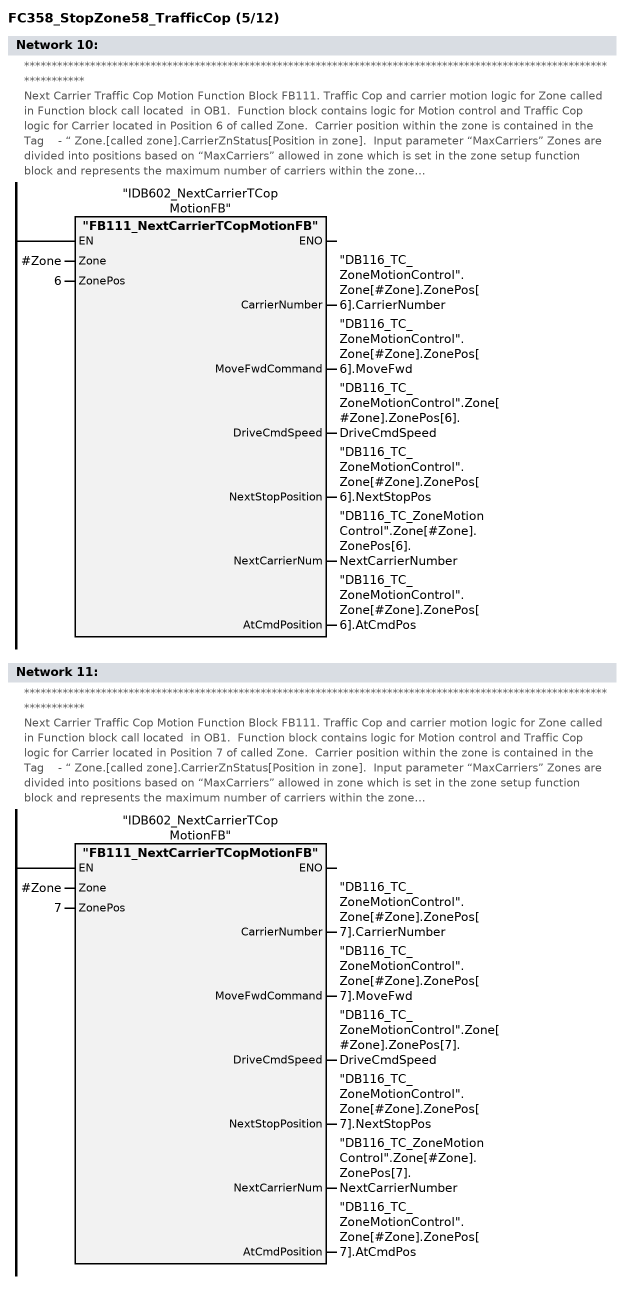
   RUNG wire#powerrail
      "IDB602_NextCarrierTCopMotionFB"(Zone := #Zone, ZonePos := 6, CarrierNumber => "DB116_TC_ZoneMotionControl".Zone[#Zone].ZonePos[6].CarrierNumber, MoveFwdCommand => "DB116_TC_ZoneMotionControl".Zone[#Zone].ZonePos[6].MoveFwd, DriveCmdSpeed => "DB116_TC_ZoneMotionControl".Zone[#Zone].ZonePos[6].DriveCmdSpeed, NextStopPosition => "DB116_TC_ZoneMotionControl".Zone[#Zone].ZonePos[6].NextStopPos, NextCarrierNum => "DB116_TC_ZoneMotionControl".Zone[#Zone].ZonePos[6].NextCarrierNumber, AtCmdPosition => "DB116_TC_ZoneMotionControl".Zone[#Zone].ZonePos[6].AtCmdPos)
   END_RUNG
   // the same network as SCL:
   "IDB602_NextCarrierTCopMotionFB"(Zone := #Zone,   // "FB111_NextCarrierTCopMotionFB"
                           ZonePos := 6,
                           CarrierNumber => "DB116_TC_ZoneMotionControl".Zone[#Zone].ZonePos[6].CarrierNumber,
                           MoveFwdCommand => "DB116_TC_ZoneMotionControl".Zone[#Zone].ZonePos[6].MoveFwd,
                           DriveCmdSpeed => "DB116_TC_ZoneMotionControl".Zone[#Zone].ZonePos[6].DriveCmdSpeed,
                           NextStopPosition => "DB116_TC_ZoneMotionControl".Zone[#Zone].ZonePos[6].NextStopPos,
                           NextCarrierNum => "DB116_TC_ZoneMotionControl".Zone[#Zone].ZonePos[6].NextCarrierNumber,
                           AtCmdPosition => "DB116_TC_ZoneMotionControl".Zone[#Zone].ZonePos[6].AtCmdPos);
END_REGION

REGION Network 11
   // *********************************************************************************************************************
   // 
   // Next Carrier Traffic Cop Motion Function Block FB111. Traffic Cop and carrier motion logic for Zone called in Function block call located  in OB1.  Function block contains logic for Motion control and Traffic Cop logic for Carrier located in Position 7 of called Zone.  Carrier position within the zone is contained in the Tag    - “ Zone.[called zone].CarrierZnStatus[Position in zone].  Input parameter “MaxCarriers” Zones are divided into positions based on “MaxCarriers” allowed in zone which is set in the zone setup function block and represents the maximum number of carriers within the zone. 
   // 
   // **********************************************************************************************************************
   RUNG wire#powerrail
      "IDB602_NextCarrierTCopMotionFB"(Zone := #Zone, ZonePos := 7, CarrierNumber => "DB116_TC_ZoneMotionControl".Zone[#Zone].ZonePos[7].CarrierNumber, MoveFwdCommand => "DB116_TC_ZoneMotionControl".Zone[#Zone].ZonePos[7].MoveFwd, DriveCmdSpeed => "DB116_TC_ZoneMotionControl".Zone[#Zone].ZonePos[7].DriveCmdSpeed, NextStopPosition => "DB116_TC_ZoneMotionControl".Zone[#Zone].ZonePos[7].NextStopPos, NextCarrierNum => "DB116_TC_ZoneMotionControl".Zone[#Zone].ZonePos[7].NextCarrierNumber, AtCmdPosition => "DB116_TC_ZoneMotionControl".Zone[#Zone].ZonePos[7].AtCmdPos)
   END_RUNG
   // the same network as SCL:
   "IDB602_NextCarrierTCopMotionFB"(Zone := #Zone,   // "FB111_NextCarrierTCopMotionFB"
                           ZonePos := 7,
                           CarrierNumber => "DB116_TC_ZoneMotionControl".Zone[#Zone].ZonePos[7].CarrierNumber,
                           MoveFwdCommand => "DB116_TC_ZoneMotionControl".Zone[#Zone].ZonePos[7].MoveFwd,
                           DriveCmdSpeed => "DB116_TC_ZoneMotionControl".Zone[#Zone].ZonePos[7].DriveCmdSpeed,
                           NextStopPosition => "DB116_TC_ZoneMotionControl".Zone[#Zone].ZonePos[7].NextStopPos,
                           NextCarrierNum => "DB116_TC_ZoneMotionControl".Zone[#Zone].ZonePos[7].NextCarrierNumber,
                           AtCmdPosition => "DB116_TC_ZoneMotionControl".Zone[#Zone].ZonePos[7].AtCmdPos);
END_REGION

REGION Network 12
   // *********************************************************************************************************************
   // 
   // Next Carrier Traffic Cop Motion Function Block FB111. Traffic Cop and carrier motion logic for Zone called in Function block call located  in OB1.  Function block contains logic for Motion control and Traffic Cop logic for Carrier located in Position 8 of called Zone.  Carrier position within the zone is contained in the Tag    - “ Zone.[called zone].CarrierZnStatus[Position in zone].  Input parameter “MaxCarriers” Zones are divided into positions based on “MaxCarriers” allowed in zone which is set in the zone setup function block and represents the maximum number of carriers within the zone. 
   // 
   // **********************************************************************************************************************
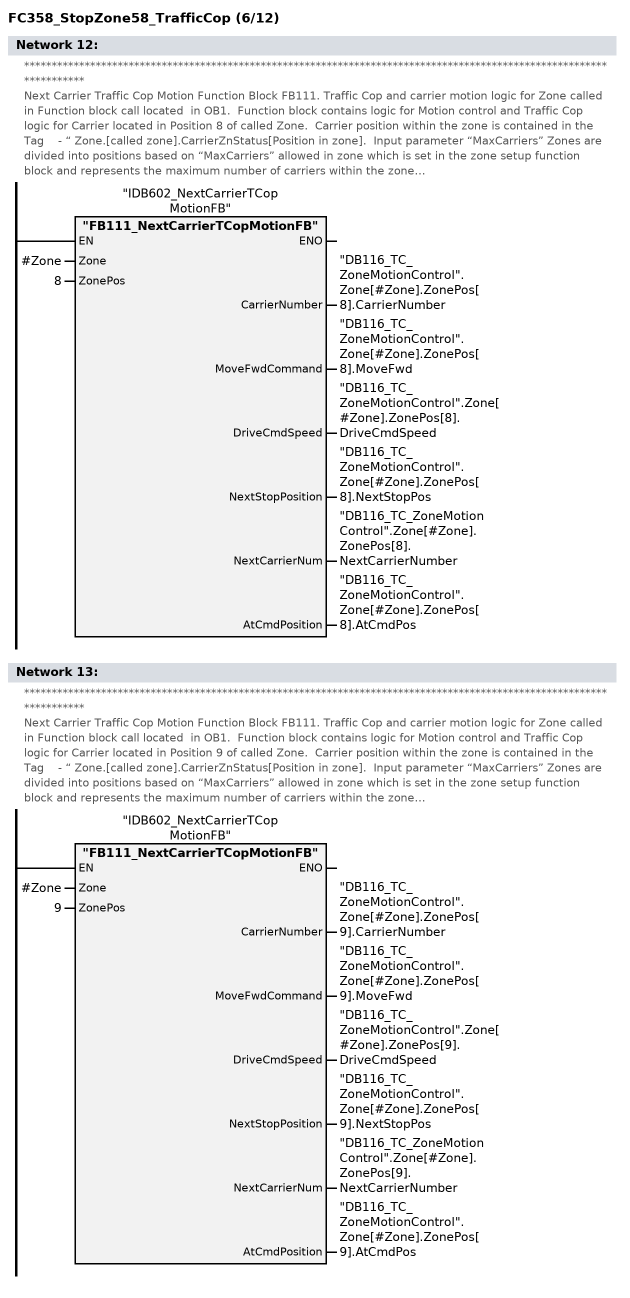
   RUNG wire#powerrail
      "IDB602_NextCarrierTCopMotionFB"(Zone := #Zone, ZonePos := 8, CarrierNumber => "DB116_TC_ZoneMotionControl".Zone[#Zone].ZonePos[8].CarrierNumber, MoveFwdCommand => "DB116_TC_ZoneMotionControl".Zone[#Zone].ZonePos[8].MoveFwd, DriveCmdSpeed => "DB116_TC_ZoneMotionControl".Zone[#Zone].ZonePos[8].DriveCmdSpeed, NextStopPosition => "DB116_TC_ZoneMotionControl".Zone[#Zone].ZonePos[8].NextStopPos, NextCarrierNum => "DB116_TC_ZoneMotionControl".Zone[#Zone].ZonePos[8].NextCarrierNumber, AtCmdPosition => "DB116_TC_ZoneMotionControl".Zone[#Zone].ZonePos[8].AtCmdPos)
   END_RUNG
   // the same network as SCL:
   "IDB602_NextCarrierTCopMotionFB"(Zone := #Zone,   // "FB111_NextCarrierTCopMotionFB"
                           ZonePos := 8,
                           CarrierNumber => "DB116_TC_ZoneMotionControl".Zone[#Zone].ZonePos[8].CarrierNumber,
                           MoveFwdCommand => "DB116_TC_ZoneMotionControl".Zone[#Zone].ZonePos[8].MoveFwd,
                           DriveCmdSpeed => "DB116_TC_ZoneMotionControl".Zone[#Zone].ZonePos[8].DriveCmdSpeed,
                           NextStopPosition => "DB116_TC_ZoneMotionControl".Zone[#Zone].ZonePos[8].NextStopPos,
                           NextCarrierNum => "DB116_TC_ZoneMotionControl".Zone[#Zone].ZonePos[8].NextCarrierNumber,
                           AtCmdPosition => "DB116_TC_ZoneMotionControl".Zone[#Zone].ZonePos[8].AtCmdPos);
END_REGION

REGION Network 13
   // *********************************************************************************************************************
   // 
   // Next Carrier Traffic Cop Motion Function Block FB111. Traffic Cop and carrier motion logic for Zone called in Function block call located  in OB1.  Function block contains logic for Motion control and Traffic Cop logic for Carrier located in Position 9 of called Zone.  Carrier position within the zone is contained in the Tag    - “ Zone.[called zone].CarrierZnStatus[Position in zone].  Input parameter “MaxCarriers” Zones are divided into positions based on “MaxCarriers” allowed in zone which is set in the zone setup function block and represents the maximum number of carriers within the zone. 
   // 
   // **********************************************************************************************************************
   RUNG wire#powerrail
      "IDB602_NextCarrierTCopMotionFB"(Zone := #Zone, ZonePos := 9, CarrierNumber => "DB116_TC_ZoneMotionControl".Zone[#Zone].ZonePos[9].CarrierNumber, MoveFwdCommand => "DB116_TC_ZoneMotionControl".Zone[#Zone].ZonePos[9].MoveFwd, DriveCmdSpeed => "DB116_TC_ZoneMotionControl".Zone[#Zone].ZonePos[9].DriveCmdSpeed, NextStopPosition => "DB116_TC_ZoneMotionControl".Zone[#Zone].ZonePos[9].NextStopPos, NextCarrierNum => "DB116_TC_ZoneMotionControl".Zone[#Zone].ZonePos[9].NextCarrierNumber, AtCmdPosition => "DB116_TC_ZoneMotionControl".Zone[#Zone].ZonePos[9].AtCmdPos)
   END_RUNG
   // the same network as SCL:
   "IDB602_NextCarrierTCopMotionFB"(Zone := #Zone,   // "FB111_NextCarrierTCopMotionFB"
                           ZonePos := 9,
                           CarrierNumber => "DB116_TC_ZoneMotionControl".Zone[#Zone].ZonePos[9].CarrierNumber,
                           MoveFwdCommand => "DB116_TC_ZoneMotionControl".Zone[#Zone].ZonePos[9].MoveFwd,
                           DriveCmdSpeed => "DB116_TC_ZoneMotionControl".Zone[#Zone].ZonePos[9].DriveCmdSpeed,
                           NextStopPosition => "DB116_TC_ZoneMotionControl".Zone[#Zone].ZonePos[9].NextStopPos,
                           NextCarrierNum => "DB116_TC_ZoneMotionControl".Zone[#Zone].ZonePos[9].NextCarrierNumber,
                           AtCmdPosition => "DB116_TC_ZoneMotionControl".Zone[#Zone].ZonePos[9].AtCmdPos);
END_REGION

REGION Network 14
   // *********************************************************************************************************************
   // 
   // Next Carrier Traffic Cop Motion Function Block FB111. Traffic Cop and carrier motion logic for Zone called in Function block call located  in OB1.  Function block contains logic for Motion control and Traffic Cop logic for Carrier located in Position 10 of called Zone.  Carrier position within the zone is contained in the Tag    - “ Zone.[called zone].CarrierZnStatus[Position in zone].  Input parameter “MaxCarriers” Zones are divided into positions based on “MaxCarriers” allowed in zone which is set in the zone setup function block and represents the maximum number of carriers within the zone. 
   // 
   // **********************************************************************************************************************
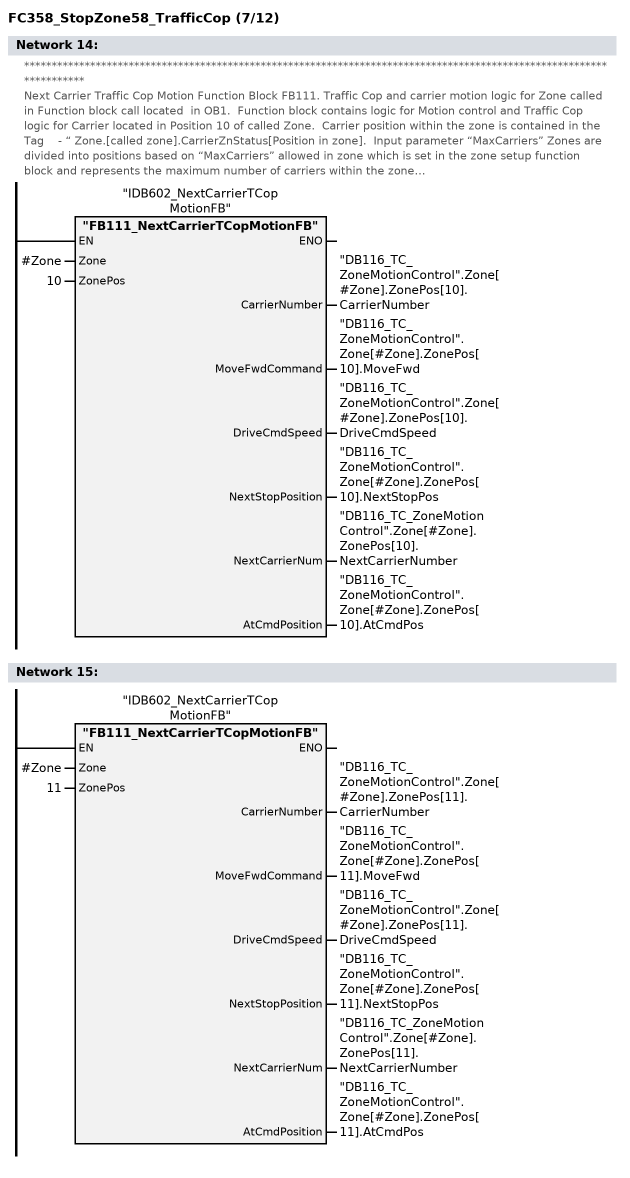
   RUNG wire#powerrail
      "IDB602_NextCarrierTCopMotionFB"(Zone := #Zone, ZonePos := 10, CarrierNumber => "DB116_TC_ZoneMotionControl".Zone[#Zone].ZonePos[10].CarrierNumber, MoveFwdCommand => "DB116_TC_ZoneMotionControl".Zone[#Zone].ZonePos[10].MoveFwd, DriveCmdSpeed => "DB116_TC_ZoneMotionControl".Zone[#Zone].ZonePos[10].DriveCmdSpeed, NextStopPosition => "DB116_TC_ZoneMotionControl".Zone[#Zone].ZonePos[10].NextStopPos, NextCarrierNum => "DB116_TC_ZoneMotionControl".Zone[#Zone].ZonePos[10].NextCarrierNumber, AtCmdPosition => "DB116_TC_ZoneMotionControl".Zone[#Zone].ZonePos[10].AtCmdPos)
   END_RUNG
   // the same network as SCL:
   "IDB602_NextCarrierTCopMotionFB"(Zone := #Zone,   // "FB111_NextCarrierTCopMotionFB"
                           ZonePos := 10,
                           CarrierNumber => "DB116_TC_ZoneMotionControl".Zone[#Zone].ZonePos[10].CarrierNumber,
                           MoveFwdCommand => "DB116_TC_ZoneMotionControl".Zone[#Zone].ZonePos[10].MoveFwd,
                           DriveCmdSpeed => "DB116_TC_ZoneMotionControl".Zone[#Zone].ZonePos[10].DriveCmdSpeed,
                           NextStopPosition => "DB116_TC_ZoneMotionControl".Zone[#Zone].ZonePos[10].NextStopPos,
                           NextCarrierNum => "DB116_TC_ZoneMotionControl".Zone[#Zone].ZonePos[10].NextCarrierNumber,
                           AtCmdPosition => "DB116_TC_ZoneMotionControl".Zone[#Zone].ZonePos[10].AtCmdPos);
END_REGION

REGION Network 15
   RUNG wire#powerrail
      "IDB602_NextCarrierTCopMotionFB"(Zone := #Zone, ZonePos := 11, CarrierNumber => "DB116_TC_ZoneMotionControl".Zone[#Zone].ZonePos[11].CarrierNumber, MoveFwdCommand => "DB116_TC_ZoneMotionControl".Zone[#Zone].ZonePos[11].MoveFwd, DriveCmdSpeed => "DB116_TC_ZoneMotionControl".Zone[#Zone].ZonePos[11].DriveCmdSpeed, NextStopPosition => "DB116_TC_ZoneMotionControl".Zone[#Zone].ZonePos[11].NextStopPos, NextCarrierNum => "DB116_TC_ZoneMotionControl".Zone[#Zone].ZonePos[11].NextCarrierNumber, AtCmdPosition => "DB116_TC_ZoneMotionControl".Zone[#Zone].ZonePos[11].AtCmdPos)
   END_RUNG
   // the same network as SCL:
   "IDB602_NextCarrierTCopMotionFB"(Zone := #Zone,   // "FB111_NextCarrierTCopMotionFB"
                           ZonePos := 11,
                           CarrierNumber => "DB116_TC_ZoneMotionControl".Zone[#Zone].ZonePos[11].CarrierNumber,
                           MoveFwdCommand => "DB116_TC_ZoneMotionControl".Zone[#Zone].ZonePos[11].MoveFwd,
                           DriveCmdSpeed => "DB116_TC_ZoneMotionControl".Zone[#Zone].ZonePos[11].DriveCmdSpeed,
                           NextStopPosition => "DB116_TC_ZoneMotionControl".Zone[#Zone].ZonePos[11].NextStopPos,
                           NextCarrierNum => "DB116_TC_ZoneMotionControl".Zone[#Zone].ZonePos[11].NextCarrierNumber,
                           AtCmdPosition => "DB116_TC_ZoneMotionControl".Zone[#Zone].ZonePos[11].AtCmdPos);
END_REGION

REGION Network 16
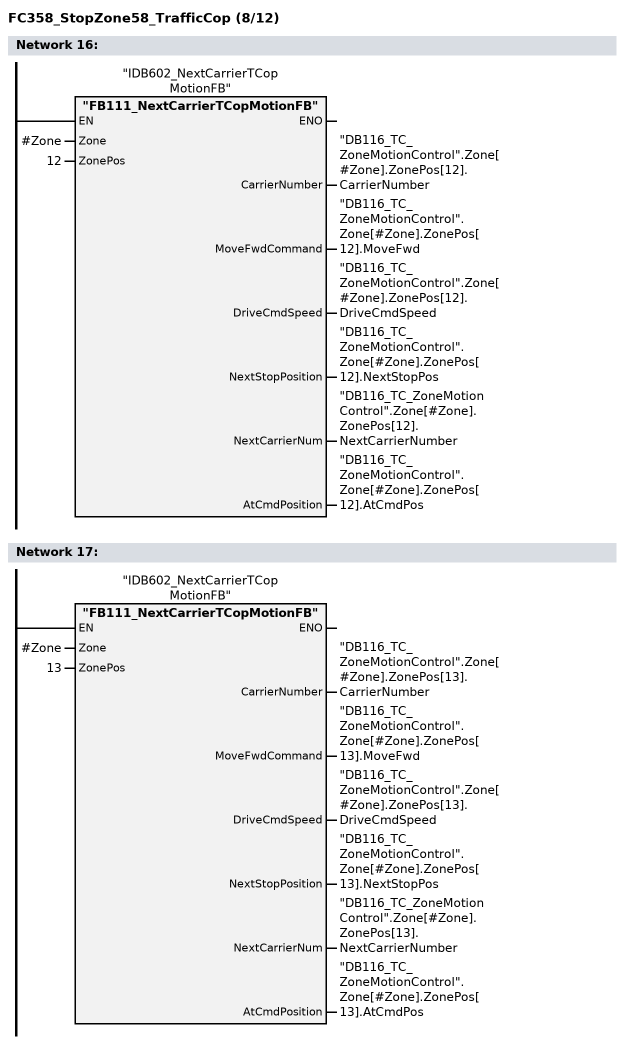
   RUNG wire#powerrail
      "IDB602_NextCarrierTCopMotionFB"(Zone := #Zone, ZonePos := 12, CarrierNumber => "DB116_TC_ZoneMotionControl".Zone[#Zone].ZonePos[12].CarrierNumber, MoveFwdCommand => "DB116_TC_ZoneMotionControl".Zone[#Zone].ZonePos[12].MoveFwd, DriveCmdSpeed => "DB116_TC_ZoneMotionControl".Zone[#Zone].ZonePos[12].DriveCmdSpeed, NextStopPosition => "DB116_TC_ZoneMotionControl".Zone[#Zone].ZonePos[12].NextStopPos, NextCarrierNum => "DB116_TC_ZoneMotionControl".Zone[#Zone].ZonePos[12].NextCarrierNumber, AtCmdPosition => "DB116_TC_ZoneMotionControl".Zone[#Zone].ZonePos[12].AtCmdPos)
   END_RUNG
   // the same network as SCL:
   "IDB602_NextCarrierTCopMotionFB"(Zone := #Zone,   // "FB111_NextCarrierTCopMotionFB"
                           ZonePos := 12,
                           CarrierNumber => "DB116_TC_ZoneMotionControl".Zone[#Zone].ZonePos[12].CarrierNumber,
                           MoveFwdCommand => "DB116_TC_ZoneMotionControl".Zone[#Zone].ZonePos[12].MoveFwd,
                           DriveCmdSpeed => "DB116_TC_ZoneMotionControl".Zone[#Zone].ZonePos[12].DriveCmdSpeed,
                           NextStopPosition => "DB116_TC_ZoneMotionControl".Zone[#Zone].ZonePos[12].NextStopPos,
                           NextCarrierNum => "DB116_TC_ZoneMotionControl".Zone[#Zone].ZonePos[12].NextCarrierNumber,
                           AtCmdPosition => "DB116_TC_ZoneMotionControl".Zone[#Zone].ZonePos[12].AtCmdPos);
END_REGION

REGION Network 17
   RUNG wire#powerrail
      "IDB602_NextCarrierTCopMotionFB"(Zone := #Zone, ZonePos := 13, CarrierNumber => "DB116_TC_ZoneMotionControl".Zone[#Zone].ZonePos[13].CarrierNumber, MoveFwdCommand => "DB116_TC_ZoneMotionControl".Zone[#Zone].ZonePos[13].MoveFwd, DriveCmdSpeed => "DB116_TC_ZoneMotionControl".Zone[#Zone].ZonePos[13].DriveCmdSpeed, NextStopPosition => "DB116_TC_ZoneMotionControl".Zone[#Zone].ZonePos[13].NextStopPos, NextCarrierNum => "DB116_TC_ZoneMotionControl".Zone[#Zone].ZonePos[13].NextCarrierNumber, AtCmdPosition => "DB116_TC_ZoneMotionControl".Zone[#Zone].ZonePos[13].AtCmdPos)
   END_RUNG
   // the same network as SCL:
   "IDB602_NextCarrierTCopMotionFB"(Zone := #Zone,   // "FB111_NextCarrierTCopMotionFB"
                           ZonePos := 13,
                           CarrierNumber => "DB116_TC_ZoneMotionControl".Zone[#Zone].ZonePos[13].CarrierNumber,
                           MoveFwdCommand => "DB116_TC_ZoneMotionControl".Zone[#Zone].ZonePos[13].MoveFwd,
                           DriveCmdSpeed => "DB116_TC_ZoneMotionControl".Zone[#Zone].ZonePos[13].DriveCmdSpeed,
                           NextStopPosition => "DB116_TC_ZoneMotionControl".Zone[#Zone].ZonePos[13].NextStopPos,
                           NextCarrierNum => "DB116_TC_ZoneMotionControl".Zone[#Zone].ZonePos[13].NextCarrierNumber,
                           AtCmdPosition => "DB116_TC_ZoneMotionControl".Zone[#Zone].ZonePos[13].AtCmdPos);
END_REGION

REGION Network 18
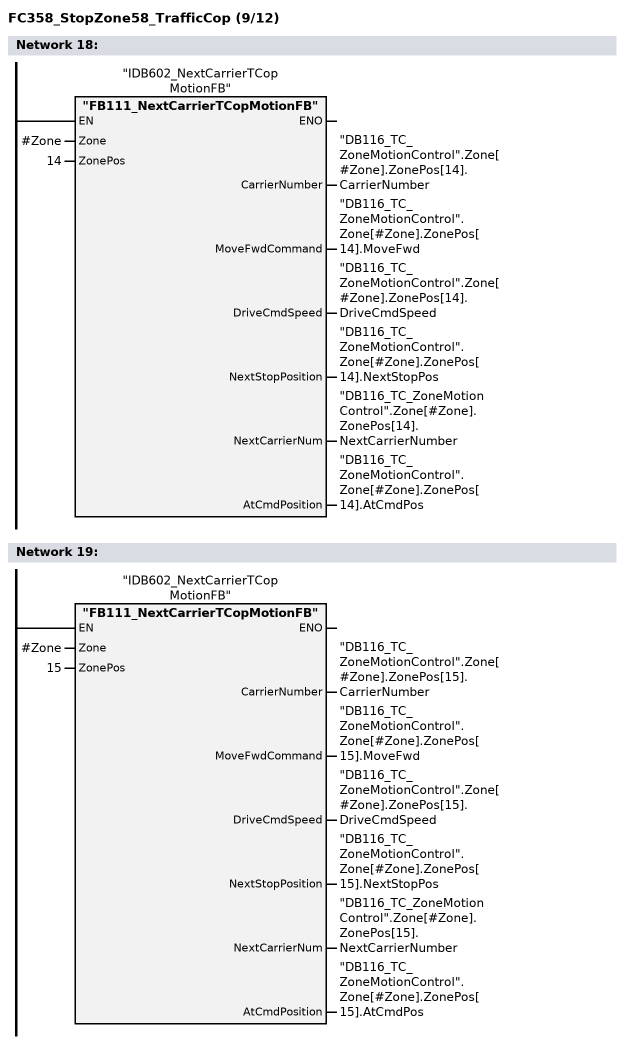
   RUNG wire#powerrail
      "IDB602_NextCarrierTCopMotionFB"(Zone := #Zone, ZonePos := 14, CarrierNumber => "DB116_TC_ZoneMotionControl".Zone[#Zone].ZonePos[14].CarrierNumber, MoveFwdCommand => "DB116_TC_ZoneMotionControl".Zone[#Zone].ZonePos[14].MoveFwd, DriveCmdSpeed => "DB116_TC_ZoneMotionControl".Zone[#Zone].ZonePos[14].DriveCmdSpeed, NextStopPosition => "DB116_TC_ZoneMotionControl".Zone[#Zone].ZonePos[14].NextStopPos, NextCarrierNum => "DB116_TC_ZoneMotionControl".Zone[#Zone].ZonePos[14].NextCarrierNumber, AtCmdPosition => "DB116_TC_ZoneMotionControl".Zone[#Zone].ZonePos[14].AtCmdPos)
   END_RUNG
   // the same network as SCL:
   "IDB602_NextCarrierTCopMotionFB"(Zone := #Zone,   // "FB111_NextCarrierTCopMotionFB"
                           ZonePos := 14,
                           CarrierNumber => "DB116_TC_ZoneMotionControl".Zone[#Zone].ZonePos[14].CarrierNumber,
                           MoveFwdCommand => "DB116_TC_ZoneMotionControl".Zone[#Zone].ZonePos[14].MoveFwd,
                           DriveCmdSpeed => "DB116_TC_ZoneMotionControl".Zone[#Zone].ZonePos[14].DriveCmdSpeed,
                           NextStopPosition => "DB116_TC_ZoneMotionControl".Zone[#Zone].ZonePos[14].NextStopPos,
                           NextCarrierNum => "DB116_TC_ZoneMotionControl".Zone[#Zone].ZonePos[14].NextCarrierNumber,
                           AtCmdPosition => "DB116_TC_ZoneMotionControl".Zone[#Zone].ZonePos[14].AtCmdPos);
END_REGION

REGION Network 19
   RUNG wire#powerrail
      "IDB602_NextCarrierTCopMotionFB"(Zone := #Zone, ZonePos := 15, CarrierNumber => "DB116_TC_ZoneMotionControl".Zone[#Zone].ZonePos[15].CarrierNumber, MoveFwdCommand => "DB116_TC_ZoneMotionControl".Zone[#Zone].ZonePos[15].MoveFwd, DriveCmdSpeed => "DB116_TC_ZoneMotionControl".Zone[#Zone].ZonePos[15].DriveCmdSpeed, NextStopPosition => "DB116_TC_ZoneMotionControl".Zone[#Zone].ZonePos[15].NextStopPos, NextCarrierNum => "DB116_TC_ZoneMotionControl".Zone[#Zone].ZonePos[15].NextCarrierNumber, AtCmdPosition => "DB116_TC_ZoneMotionControl".Zone[#Zone].ZonePos[15].AtCmdPos)
   END_RUNG
   // the same network as SCL:
   "IDB602_NextCarrierTCopMotionFB"(Zone := #Zone,   // "FB111_NextCarrierTCopMotionFB"
                           ZonePos := 15,
                           CarrierNumber => "DB116_TC_ZoneMotionControl".Zone[#Zone].ZonePos[15].CarrierNumber,
                           MoveFwdCommand => "DB116_TC_ZoneMotionControl".Zone[#Zone].ZonePos[15].MoveFwd,
                           DriveCmdSpeed => "DB116_TC_ZoneMotionControl".Zone[#Zone].ZonePos[15].DriveCmdSpeed,
                           NextStopPosition => "DB116_TC_ZoneMotionControl".Zone[#Zone].ZonePos[15].NextStopPos,
                           NextCarrierNum => "DB116_TC_ZoneMotionControl".Zone[#Zone].ZonePos[15].NextCarrierNumber,
                           AtCmdPosition => "DB116_TC_ZoneMotionControl".Zone[#Zone].ZonePos[15].AtCmdPos);
END_REGION

REGION Network 20
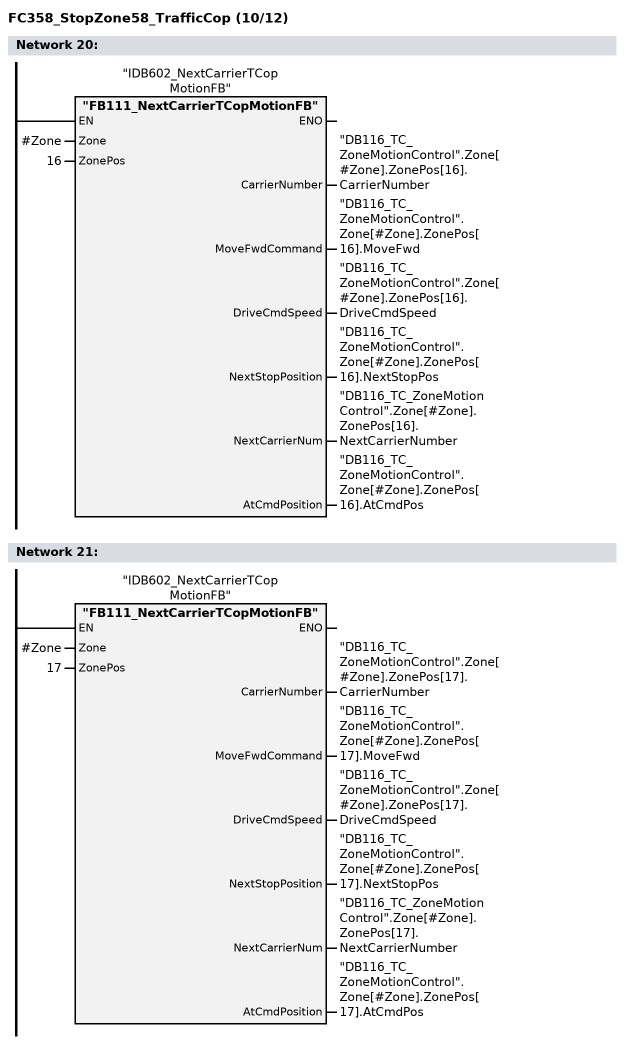
   RUNG wire#powerrail
      "IDB602_NextCarrierTCopMotionFB"(Zone := #Zone, ZonePos := 16, CarrierNumber => "DB116_TC_ZoneMotionControl".Zone[#Zone].ZonePos[16].CarrierNumber, MoveFwdCommand => "DB116_TC_ZoneMotionControl".Zone[#Zone].ZonePos[16].MoveFwd, DriveCmdSpeed => "DB116_TC_ZoneMotionControl".Zone[#Zone].ZonePos[16].DriveCmdSpeed, NextStopPosition => "DB116_TC_ZoneMotionControl".Zone[#Zone].ZonePos[16].NextStopPos, NextCarrierNum => "DB116_TC_ZoneMotionControl".Zone[#Zone].ZonePos[16].NextCarrierNumber, AtCmdPosition => "DB116_TC_ZoneMotionControl".Zone[#Zone].ZonePos[16].AtCmdPos)
   END_RUNG
   // the same network as SCL:
   "IDB602_NextCarrierTCopMotionFB"(Zone := #Zone,   // "FB111_NextCarrierTCopMotionFB"
                           ZonePos := 16,
                           CarrierNumber => "DB116_TC_ZoneMotionControl".Zone[#Zone].ZonePos[16].CarrierNumber,
                           MoveFwdCommand => "DB116_TC_ZoneMotionControl".Zone[#Zone].ZonePos[16].MoveFwd,
                           DriveCmdSpeed => "DB116_TC_ZoneMotionControl".Zone[#Zone].ZonePos[16].DriveCmdSpeed,
                           NextStopPosition => "DB116_TC_ZoneMotionControl".Zone[#Zone].ZonePos[16].NextStopPos,
                           NextCarrierNum => "DB116_TC_ZoneMotionControl".Zone[#Zone].ZonePos[16].NextCarrierNumber,
                           AtCmdPosition => "DB116_TC_ZoneMotionControl".Zone[#Zone].ZonePos[16].AtCmdPos);
END_REGION

REGION Network 21
   RUNG wire#powerrail
      "IDB602_NextCarrierTCopMotionFB"(Zone := #Zone, ZonePos := 17, CarrierNumber => "DB116_TC_ZoneMotionControl".Zone[#Zone].ZonePos[17].CarrierNumber, MoveFwdCommand => "DB116_TC_ZoneMotionControl".Zone[#Zone].ZonePos[17].MoveFwd, DriveCmdSpeed => "DB116_TC_ZoneMotionControl".Zone[#Zone].ZonePos[17].DriveCmdSpeed, NextStopPosition => "DB116_TC_ZoneMotionControl".Zone[#Zone].ZonePos[17].NextStopPos, NextCarrierNum => "DB116_TC_ZoneMotionControl".Zone[#Zone].ZonePos[17].NextCarrierNumber, AtCmdPosition => "DB116_TC_ZoneMotionControl".Zone[#Zone].ZonePos[17].AtCmdPos)
   END_RUNG
   // the same network as SCL:
   "IDB602_NextCarrierTCopMotionFB"(Zone := #Zone,   // "FB111_NextCarrierTCopMotionFB"
                           ZonePos := 17,
                           CarrierNumber => "DB116_TC_ZoneMotionControl".Zone[#Zone].ZonePos[17].CarrierNumber,
                           MoveFwdCommand => "DB116_TC_ZoneMotionControl".Zone[#Zone].ZonePos[17].MoveFwd,
                           DriveCmdSpeed => "DB116_TC_ZoneMotionControl".Zone[#Zone].ZonePos[17].DriveCmdSpeed,
                           NextStopPosition => "DB116_TC_ZoneMotionControl".Zone[#Zone].ZonePos[17].NextStopPos,
                           NextCarrierNum => "DB116_TC_ZoneMotionControl".Zone[#Zone].ZonePos[17].NextCarrierNumber,
                           AtCmdPosition => "DB116_TC_ZoneMotionControl".Zone[#Zone].ZonePos[17].AtCmdPos);
END_REGION

REGION Network 22
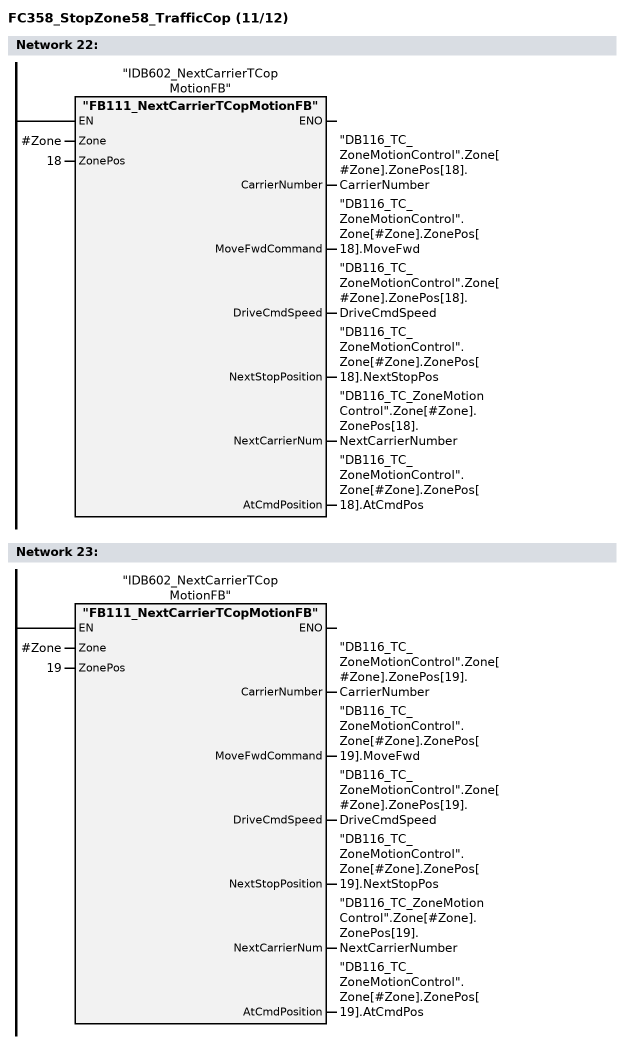
   RUNG wire#powerrail
      "IDB602_NextCarrierTCopMotionFB"(Zone := #Zone, ZonePos := 18, CarrierNumber => "DB116_TC_ZoneMotionControl".Zone[#Zone].ZonePos[18].CarrierNumber, MoveFwdCommand => "DB116_TC_ZoneMotionControl".Zone[#Zone].ZonePos[18].MoveFwd, DriveCmdSpeed => "DB116_TC_ZoneMotionControl".Zone[#Zone].ZonePos[18].DriveCmdSpeed, NextStopPosition => "DB116_TC_ZoneMotionControl".Zone[#Zone].ZonePos[18].NextStopPos, NextCarrierNum => "DB116_TC_ZoneMotionControl".Zone[#Zone].ZonePos[18].NextCarrierNumber, AtCmdPosition => "DB116_TC_ZoneMotionControl".Zone[#Zone].ZonePos[18].AtCmdPos)
   END_RUNG
   // the same network as SCL:
   "IDB602_NextCarrierTCopMotionFB"(Zone := #Zone,   // "FB111_NextCarrierTCopMotionFB"
                           ZonePos := 18,
                           CarrierNumber => "DB116_TC_ZoneMotionControl".Zone[#Zone].ZonePos[18].CarrierNumber,
                           MoveFwdCommand => "DB116_TC_ZoneMotionControl".Zone[#Zone].ZonePos[18].MoveFwd,
                           DriveCmdSpeed => "DB116_TC_ZoneMotionControl".Zone[#Zone].ZonePos[18].DriveCmdSpeed,
                           NextStopPosition => "DB116_TC_ZoneMotionControl".Zone[#Zone].ZonePos[18].NextStopPos,
                           NextCarrierNum => "DB116_TC_ZoneMotionControl".Zone[#Zone].ZonePos[18].NextCarrierNumber,
                           AtCmdPosition => "DB116_TC_ZoneMotionControl".Zone[#Zone].ZonePos[18].AtCmdPos);
END_REGION

REGION Network 23
   RUNG wire#powerrail
      "IDB602_NextCarrierTCopMotionFB"(Zone := #Zone, ZonePos := 19, CarrierNumber => "DB116_TC_ZoneMotionControl".Zone[#Zone].ZonePos[19].CarrierNumber, MoveFwdCommand => "DB116_TC_ZoneMotionControl".Zone[#Zone].ZonePos[19].MoveFwd, DriveCmdSpeed => "DB116_TC_ZoneMotionControl".Zone[#Zone].ZonePos[19].DriveCmdSpeed, NextStopPosition => "DB116_TC_ZoneMotionControl".Zone[#Zone].ZonePos[19].NextStopPos, NextCarrierNum => "DB116_TC_ZoneMotionControl".Zone[#Zone].ZonePos[19].NextCarrierNumber, AtCmdPosition => "DB116_TC_ZoneMotionControl".Zone[#Zone].ZonePos[19].AtCmdPos)
   END_RUNG
   // the same network as SCL:
   "IDB602_NextCarrierTCopMotionFB"(Zone := #Zone,   // "FB111_NextCarrierTCopMotionFB"
                           ZonePos := 19,
                           CarrierNumber => "DB116_TC_ZoneMotionControl".Zone[#Zone].ZonePos[19].CarrierNumber,
                           MoveFwdCommand => "DB116_TC_ZoneMotionControl".Zone[#Zone].ZonePos[19].MoveFwd,
                           DriveCmdSpeed => "DB116_TC_ZoneMotionControl".Zone[#Zone].ZonePos[19].DriveCmdSpeed,
                           NextStopPosition => "DB116_TC_ZoneMotionControl".Zone[#Zone].ZonePos[19].NextStopPos,
                           NextCarrierNum => "DB116_TC_ZoneMotionControl".Zone[#Zone].ZonePos[19].NextCarrierNumber,
                           AtCmdPosition => "DB116_TC_ZoneMotionControl".Zone[#Zone].ZonePos[19].AtCmdPos);
END_REGION

REGION Network 24
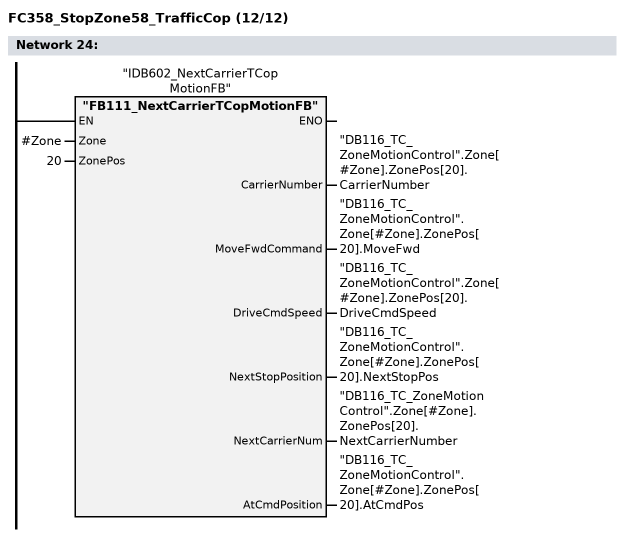
   RUNG wire#powerrail
      "IDB602_NextCarrierTCopMotionFB"(Zone := #Zone, ZonePos := 20, CarrierNumber => "DB116_TC_ZoneMotionControl".Zone[#Zone].ZonePos[20].CarrierNumber, MoveFwdCommand => "DB116_TC_ZoneMotionControl".Zone[#Zone].ZonePos[20].MoveFwd, DriveCmdSpeed => "DB116_TC_ZoneMotionControl".Zone[#Zone].ZonePos[20].DriveCmdSpeed, NextStopPosition => "DB116_TC_ZoneMotionControl".Zone[#Zone].ZonePos[20].NextStopPos, NextCarrierNum => "DB116_TC_ZoneMotionControl".Zone[#Zone].ZonePos[20].NextCarrierNumber, AtCmdPosition => "DB116_TC_ZoneMotionControl".Zone[#Zone].ZonePos[20].AtCmdPos)
   END_RUNG
   // the same network as SCL:
   "IDB602_NextCarrierTCopMotionFB"(Zone := #Zone,   // "FB111_NextCarrierTCopMotionFB"
                           ZonePos := 20,
                           CarrierNumber => "DB116_TC_ZoneMotionControl".Zone[#Zone].ZonePos[20].CarrierNumber,
                           MoveFwdCommand => "DB116_TC_ZoneMotionControl".Zone[#Zone].ZonePos[20].MoveFwd,
                           DriveCmdSpeed => "DB116_TC_ZoneMotionControl".Zone[#Zone].ZonePos[20].DriveCmdSpeed,
                           NextStopPosition => "DB116_TC_ZoneMotionControl".Zone[#Zone].ZonePos[20].NextStopPos,
                           NextCarrierNum => "DB116_TC_ZoneMotionControl".Zone[#Zone].ZonePos[20].NextCarrierNumber,
                           AtCmdPosition => "DB116_TC_ZoneMotionControl".Zone[#Zone].ZonePos[20].AtCmdPos);
END_REGION
END_FUNCTION

FUNCTION "FC400_HMI_Status" : Void   // FC400, LAD
{ S7_Optimized_Access := 'TRUE' }
VERSION : 0.1
BEGIN

REGION Network 1
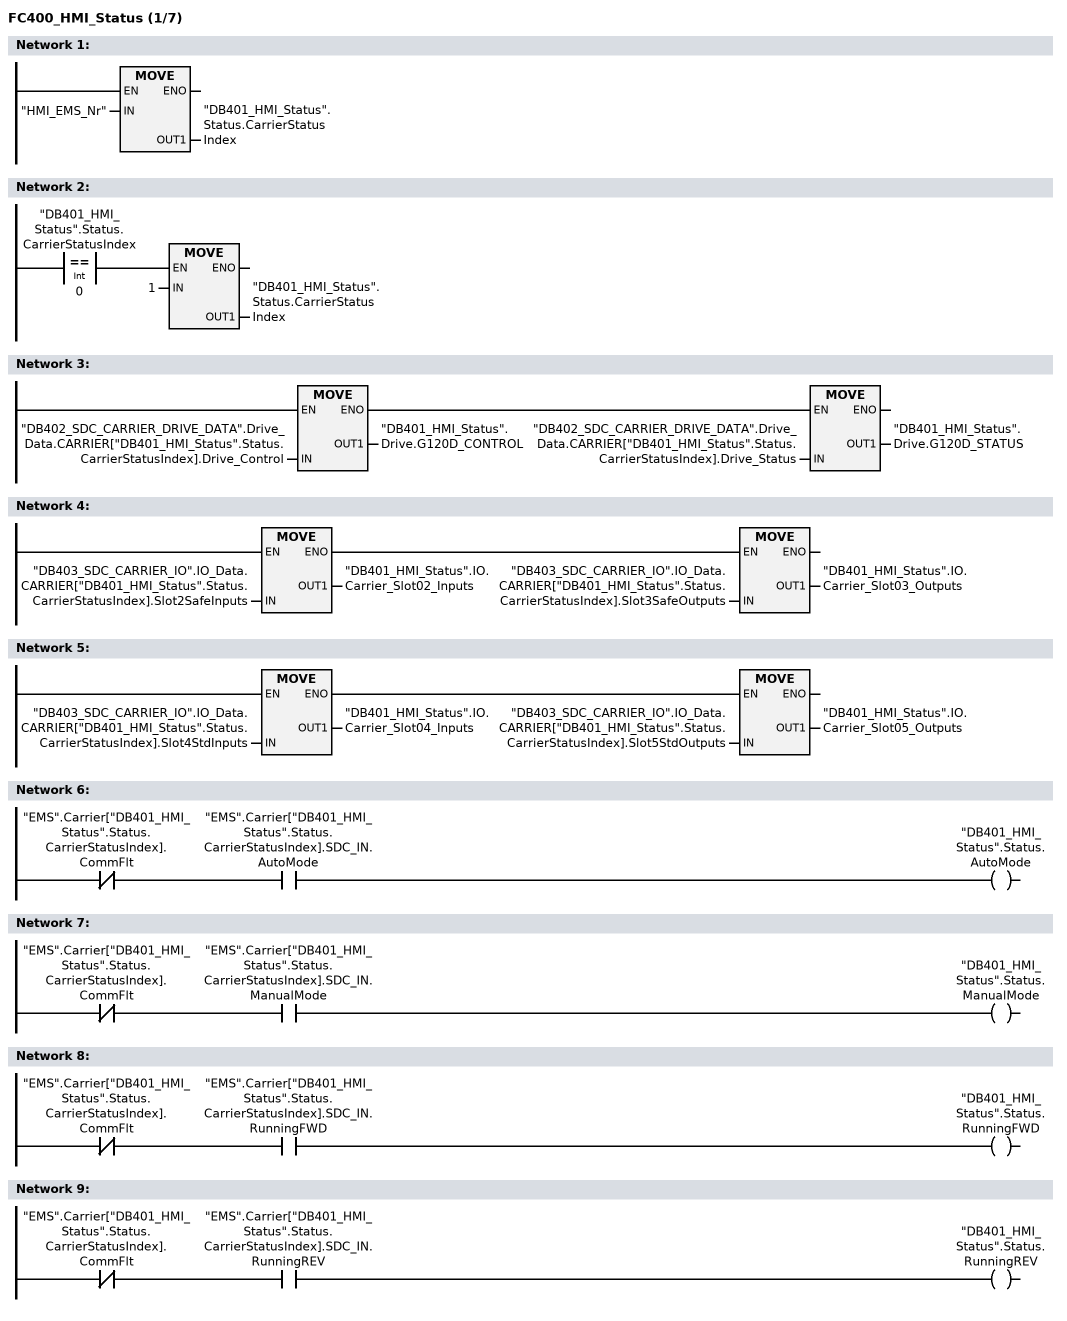
   RUNG wire#powerrail
      Move(in := "HMI_EMS_Nr", out1 => "DB401_HMI_Status".Status.CarrierStatusIndex)
   END_RUNG
   // the same network as SCL:
   "DB401_HMI_Status".Status.CarrierStatusIndex := "HMI_EMS_Nr";
END_REGION

REGION Network 2
   RUNG wire#powerrail
      { S7_Templates := "SrcType := Int" } EQ_Contact(in1 := "DB401_HMI_Status".Status.CarrierStatusIndex, in2 := 0)
      Move(in := 1, out1 => "DB401_HMI_Status".Status.CarrierStatusIndex)
   END_RUNG
   // the same network as SCL:
   IF "DB401_HMI_Status".Status.CarrierStatusIndex = 0 THEN
       "DB401_HMI_Status".Status.CarrierStatusIndex := 1;
   END_IF;
END_REGION

REGION Network 3
   RUNG wire#powerrail
      Move(in := "DB402_SDC_CARRIER_DRIVE_DATA".Drive_Data.CARRIER["DB401_HMI_Status".Status.CarrierStatusIndex].Drive_Control, out1 => "DB401_HMI_Status".Drive.G120D_CONTROL)
      Move(in := "DB402_SDC_CARRIER_DRIVE_DATA".Drive_Data.CARRIER["DB401_HMI_Status".Status.CarrierStatusIndex].Drive_Status, out1 => "DB401_HMI_Status".Drive.G120D_STATUS)
   END_RUNG
   // the same network as SCL:
   "DB401_HMI_Status".Drive.G120D_CONTROL := "DB402_SDC_CARRIER_DRIVE_DATA".Drive_Data.CARRIER["DB401_HMI_Status".Status.CarrierStatusIndex].Drive_Control;
   "DB401_HMI_Status".Drive.G120D_STATUS := "DB402_SDC_CARRIER_DRIVE_DATA".Drive_Data.CARRIER["DB401_HMI_Status".Status.CarrierStatusIndex].Drive_Status;
END_REGION

REGION Network 4
   RUNG wire#powerrail
      Move(in := "DB403_SDC_CARRIER_IO".IO_Data.CARRIER["DB401_HMI_Status".Status.CarrierStatusIndex].Slot2SafeInputs, out1 => "DB401_HMI_Status".IO.Carrier_Slot02_Inputs)
      Move(in := "DB403_SDC_CARRIER_IO".IO_Data.CARRIER["DB401_HMI_Status".Status.CarrierStatusIndex].Slot3SafeOutputs, out1 => "DB401_HMI_Status".IO.Carrier_Slot03_Outputs)
   END_RUNG
   // the same network as SCL:
   "DB401_HMI_Status".IO.Carrier_Slot02_Inputs := "DB403_SDC_CARRIER_IO".IO_Data.CARRIER["DB401_HMI_Status".Status.CarrierStatusIndex].Slot2SafeInputs;
   "DB401_HMI_Status".IO.Carrier_Slot03_Outputs := "DB403_SDC_CARRIER_IO".IO_Data.CARRIER["DB401_HMI_Status".Status.CarrierStatusIndex].Slot3SafeOutputs;
END_REGION

REGION Network 5
   RUNG wire#powerrail
      Move(in := "DB403_SDC_CARRIER_IO".IO_Data.CARRIER["DB401_HMI_Status".Status.CarrierStatusIndex].Slot4StdInputs, out1 => "DB401_HMI_Status".IO.Carrier_Slot04_Inputs)
      Move(in := "DB403_SDC_CARRIER_IO".IO_Data.CARRIER["DB401_HMI_Status".Status.CarrierStatusIndex].Slot5StdOutputs, out1 => "DB401_HMI_Status".IO.Carrier_Slot05_Outputs)
   END_RUNG
   // the same network as SCL:
   "DB401_HMI_Status".IO.Carrier_Slot04_Inputs := "DB403_SDC_CARRIER_IO".IO_Data.CARRIER["DB401_HMI_Status".Status.CarrierStatusIndex].Slot4StdInputs;
   "DB401_HMI_Status".IO.Carrier_Slot05_Outputs := "DB403_SDC_CARRIER_IO".IO_Data.CARRIER["DB401_HMI_Status".Status.CarrierStatusIndex].Slot5StdOutputs;
END_REGION

REGION Network 6
   RUNG wire#powerrail
      I_Contact( "EMS".Carrier["DB401_HMI_Status".Status.CarrierStatusIndex].CommFlt )
      Contact( "EMS".Carrier["DB401_HMI_Status".Status.CarrierStatusIndex].SDC_IN.AutoMode )
      Coil( "DB401_HMI_Status".Status.AutoMode )
   END_RUNG
   // the same network as SCL:
   "DB401_HMI_Status".Status.AutoMode := NOT "EMS".Carrier["DB401_HMI_Status".Status.CarrierStatusIndex].CommFlt AND "EMS".Carrier["DB401_HMI_Status".Status.CarrierStatusIndex].SDC_IN.AutoMode;
END_REGION

REGION Network 7
   RUNG wire#powerrail
      I_Contact( "EMS".Carrier["DB401_HMI_Status".Status.CarrierStatusIndex].CommFlt )
      Contact( "EMS".Carrier["DB401_HMI_Status".Status.CarrierStatusIndex].SDC_IN.ManualMode )
      Coil( "DB401_HMI_Status".Status.ManualMode )
   END_RUNG
   // the same network as SCL:
   "DB401_HMI_Status".Status.ManualMode := NOT "EMS".Carrier["DB401_HMI_Status".Status.CarrierStatusIndex].CommFlt AND "EMS".Carrier["DB401_HMI_Status".Status.CarrierStatusIndex].SDC_IN.ManualMode;
END_REGION

REGION Network 8
   RUNG wire#powerrail
      I_Contact( "EMS".Carrier["DB401_HMI_Status".Status.CarrierStatusIndex].CommFlt )
      Contact( "EMS".Carrier["DB401_HMI_Status".Status.CarrierStatusIndex].SDC_IN.RunningFWD )
      Coil( "DB401_HMI_Status".Status.RunningFWD )
   END_RUNG
   // the same network as SCL:
   "DB401_HMI_Status".Status.RunningFWD := NOT "EMS".Carrier["DB401_HMI_Status".Status.CarrierStatusIndex].CommFlt AND "EMS".Carrier["DB401_HMI_Status".Status.CarrierStatusIndex].SDC_IN.RunningFWD;
END_REGION
